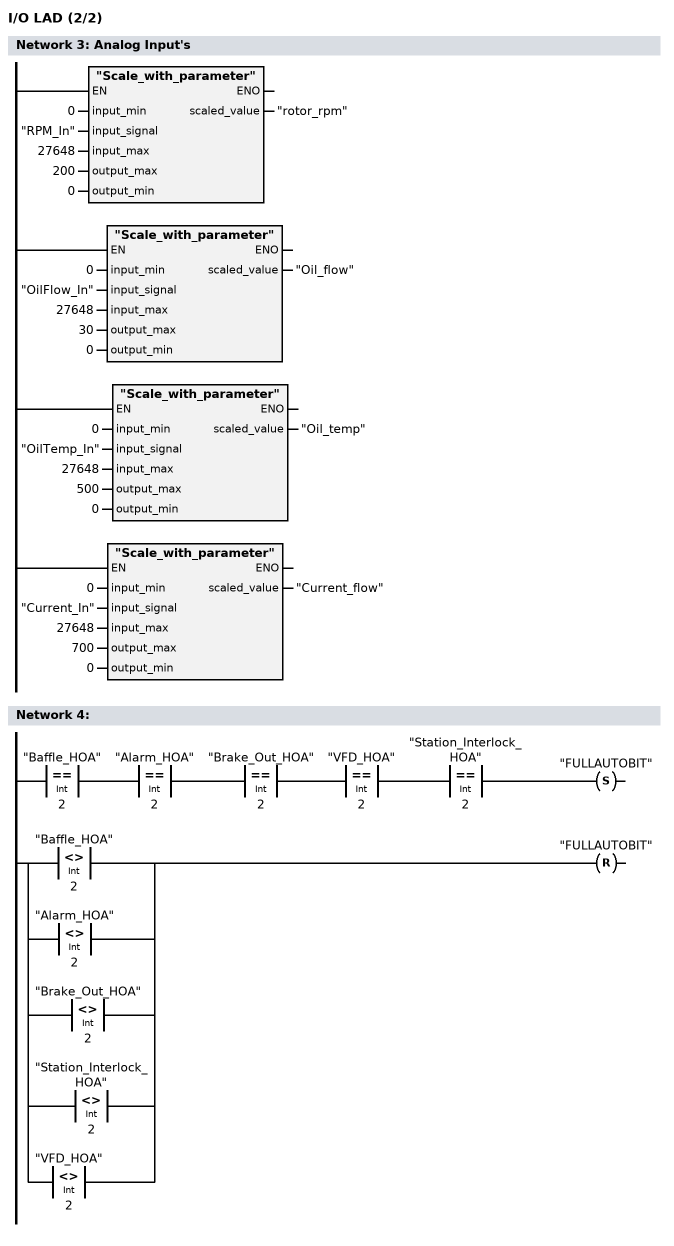
   RUNG wire#powerrail
      "Scale_with_parameter"(input_min := 0, input_signal := "RPM_In", input_max := 27648, output_max := 200, output_min := 0, scaled_value => "rotor_rpm")
   END_RUNG
   RUNG wire#powerrail
      "Scale_with_parameter"(input_min := 0, input_signal := "OilFlow_In", input_max := 27648, output_max := 30, output_min := 0, scaled_value => "Oil_flow")
   END_RUNG
   RUNG wire#powerrail
      "Scale_with_parameter"(input_min := 0, input_signal := "OilTemp_In", input_max := 27648, output_max := 500, output_min := 0, scaled_value => "Oil_temp")
   END_RUNG
   RUNG wire#powerrail
      "Scale_with_parameter"(input_min := 0, input_signal := "Current_In", input_max := 27648, output_max := 700, output_min := 0, scaled_value => "Current_flow")
   END_RUNG
   // the same network as SCL:
   "Scale_with_parameter"(input_min := 0,
                          input_signal := "RPM_In",
                          input_max := 27648,
                          output_max := 200,
                          output_min := 0,
                          scaled_value => "rotor_rpm");
   "Scale_with_parameter"(input_min := 0,
                          input_signal := "OilFlow_In",
                          input_max := 27648,
                          output_max := 30,
                          output_min := 0,
                          scaled_value => "Oil_flow");
   "Scale_with_parameter"(input_min := 0,
                          input_signal := "OilTemp_In",
                          input_max := 27648,
                          output_max := 500,
                          output_min := 0,
                          scaled_value => "Oil_temp");
   "Scale_with_parameter"(input_min := 0,
                          input_signal := "Current_In",
                          input_max := 27648,
                          output_max := 700,
                          output_min := 0,
                          scaled_value => "Current_flow");
END_REGION

REGION Network 4
   RUNG wire#powerrail
      { S7_Templates := "SrcType := Int" } EQ_Contact(in1 := "Baffle_HOA", in2 := 2)
      { S7_Templates := "SrcType := Int" } EQ_Contact(in1 := "Alarm_HOA", in2 := 2)
      { S7_Templates := "SrcType := Int" } EQ_Contact(in1 := "Brake_Out_HOA", in2 := 2)
      { S7_Templates := "SrcType := Int" } EQ_Contact(in1 := "VFD_HOA", in2 := 2)
      { S7_Templates := "SrcType := Int" } EQ_Contact(in1 := "Station_Interlock_HOA", in2 := 2)
      S_Coil( "FULLAUTOBIT" )
   END_RUNG
   RUNG wire#powerrail
      { S7_Templates := "SrcType := Int" } NE_Contact(in1 := "Baffle_HOA", in2 := 2)
      wire#w1
      R_Coil( "FULLAUTOBIT" )
   END_RUNG
   RUNG wire#powerrail
      { S7_Templates := "SrcType := Int" } NE_Contact(in1 := "Alarm_HOA", in2 := 2)
   END_RUNG wire#w1
   RUNG wire#powerrail
      { S7_Templates := "SrcType := Int" } NE_Contact(in1 := "Brake_Out_HOA", in2 := 2)
   END_RUNG wire#w1
   RUNG wire#powerrail
      { S7_Templates := "SrcType := Int" } NE_Contact(in1 := "Station_Interlock_HOA", in2 := 2)
   END_RUNG wire#w1
   RUNG wire#powerrail
      { S7_Templates := "SrcType := Int" } NE_Contact(in1 := "VFD_HOA", in2 := 2)
   END_RUNG wire#w1
   // the same network as SCL:
   IF ("Baffle_HOA" = 2) AND ("Alarm_HOA" = 2) AND ("Brake_Out_HOA" = 2) AND ("VFD_HOA" = 2) AND ("Station_Interlock_HOA" = 2) THEN
       "FULLAUTOBIT" := TRUE;
   END_IF;
   IF ("Baffle_HOA" <> 2) OR ("Alarm_HOA" <> 2) OR ("Brake_Out_HOA" <> 2) OR ("Station_Interlock_HOA" <> 2) OR ("VFD_HOA" <> 2) THEN
       "FULLAUTOBIT" := FALSE;
   END_IF;
END_REGION
END_FUNCTION_BLOCK

FUNCTION_BLOCK "HOA_LAD"   // FB6, LAD
TITLE = Push Button for HOA (OFF, HAND, AUTO)
{ S7_Optimized_Access := 'TRUE' }
VERSION : 0.1
   VAR
      Os3 : Bool;
      Os2 : Bool;
      Os1 : Bool;
      Os4 : Bool;
      Os5 : Bool;
      Os6 : Bool;
      Os7 : Bool;
      Os8 : Bool;
      Os9 : Bool;
      Os10 : Bool;
      Os11 : Bool;
      Os12 : Bool;
   END_VAR
   VAR_TEMP   // added for the SCL form of the ladder/FBD networks
      _w1 : Bool;
      _w2 : Bool;
      _w3 : Bool;
   END_VAR
BEGIN

REGION Network 1
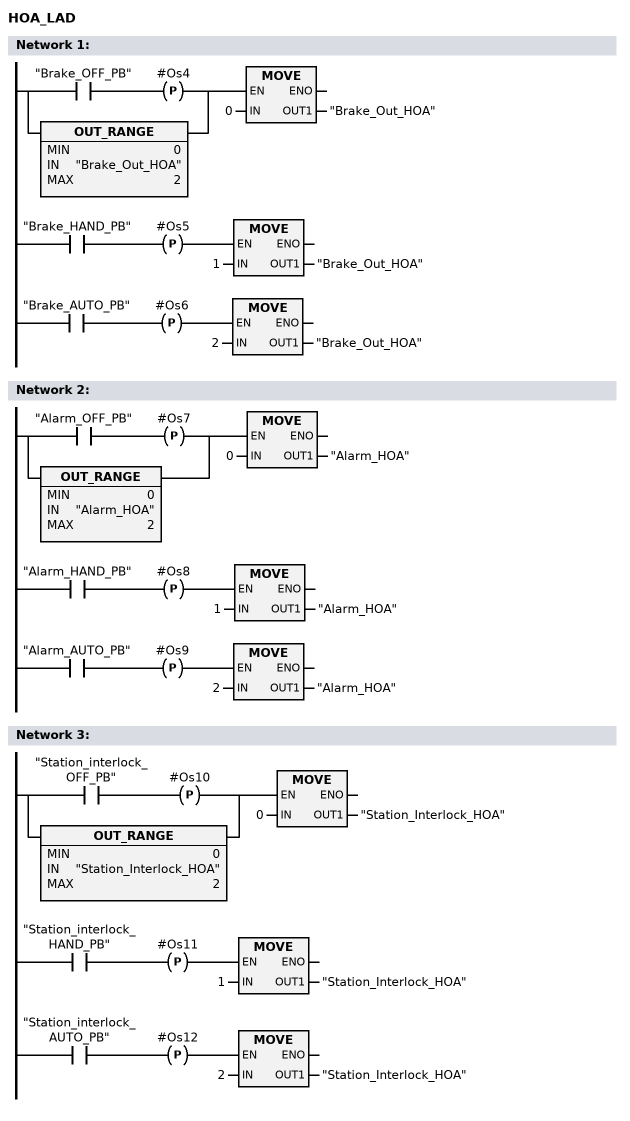
   #_w1 := "Brake_OFF_PB" AND NOT #Os4;   // rising edge
   #Os4 := "Brake_OFF_PB";
   IF #_w1 OR ("Brake_Out_HOA" < 0) OR ("Brake_Out_HOA" > 2) THEN "Brake_Out_HOA" := 0; END_IF;
   #_w2 := "Brake_HAND_PB" AND NOT #Os5;   // rising edge
   #Os5 := "Brake_HAND_PB";
   IF #_w2 THEN "Brake_Out_HOA" := 1; END_IF;
   #_w3 := "Brake_AUTO_PB" AND NOT #Os6;   // rising edge
   #Os6 := "Brake_AUTO_PB";
   IF #_w3 THEN "Brake_Out_HOA" := 2; END_IF;
END_REGION

REGION Network 2
   #_w1 := "Alarm_OFF_PB" AND NOT #Os7;   // rising edge
   #Os7 := "Alarm_OFF_PB";
   IF #_w1 OR ("Alarm_HOA" < 0) OR ("Alarm_HOA" > 2) THEN "Alarm_HOA" := 0; END_IF;
   #_w2 := "Alarm_HAND_PB" AND NOT #Os8;   // rising edge
   #Os8 := "Alarm_HAND_PB";
   IF #_w2 THEN "Alarm_HOA" := 1; END_IF;
   #_w3 := "Alarm_AUTO_PB" AND NOT #Os9;   // rising edge
   #Os9 := "Alarm_AUTO_PB";
   IF #_w3 THEN "Alarm_HOA" := 2; END_IF;
END_REGION

REGION Network 3
   #_w1 := "Station_interlock_OFF_PB" AND NOT #Os10;   // rising edge
   #Os10 := "Station_interlock_OFF_PB";
   IF #_w1 OR ("Station_Interlock_HOA" < 0) OR ("Station_Interlock_HOA" > 2) THEN
       "Station_Interlock_HOA" := 0;
   END_IF;
   #_w2 := "Station_interlock_HAND_PB" AND NOT #Os11;   // rising edge
   #Os11 := "Station_interlock_HAND_PB";
   IF #_w2 THEN "Station_Interlock_HOA" := 1; END_IF;
   #_w3 := "Station_interlock_AUTO_PB" AND NOT #Os12;   // rising edge
   #Os12 := "Station_interlock_AUTO_PB";
   IF #_w3 THEN "Station_Interlock_HOA" := 2; END_IF;
END_REGION
END_FUNCTION_BLOCK

FUNCTION_BLOCK "Alarm_LAD"   // FB10, LAD
{ S7_Optimized_Access := 'TRUE' }
VERSION : 0.1
   VAR
      OS1 : Bool;
      OS2 : Bool;
      OS3 : Bool;
      OS4 : Bool;
      OS5 : Bool;
      OS6 : Bool;
      OS7 : Bool;
      os8 : Bool;
   END_VAR
   VAR_TEMP
      tp1 : Int;
      OLFD : Time;
      OFL_AT : Bool;
      tp2 : Int;
      OCD : Time;
      OC_AT : Bool;
      tp3 : Int;
      HOT : Time;
      HOT_AT : Bool;
      tp4 : Int;
      ROS : Time;
      ROS_AT : Bool;
      tp5 : Int;
      OHF : Time;
      OHF_AT : Bool;
      tp6 : Int;
      BF : Time;
      BF_AT : Bool;
      ES_AT : Bool;
      AlarmTrigger : Bool;
   END_VAR
   VAR_TEMP   // added for the SCL form of the ladder/FBD networks
      _w1 : Bool;
      _w2 : Bool;
   END_VAR
BEGIN

REGION Network 1: Alarm for OIL LOW FLOW
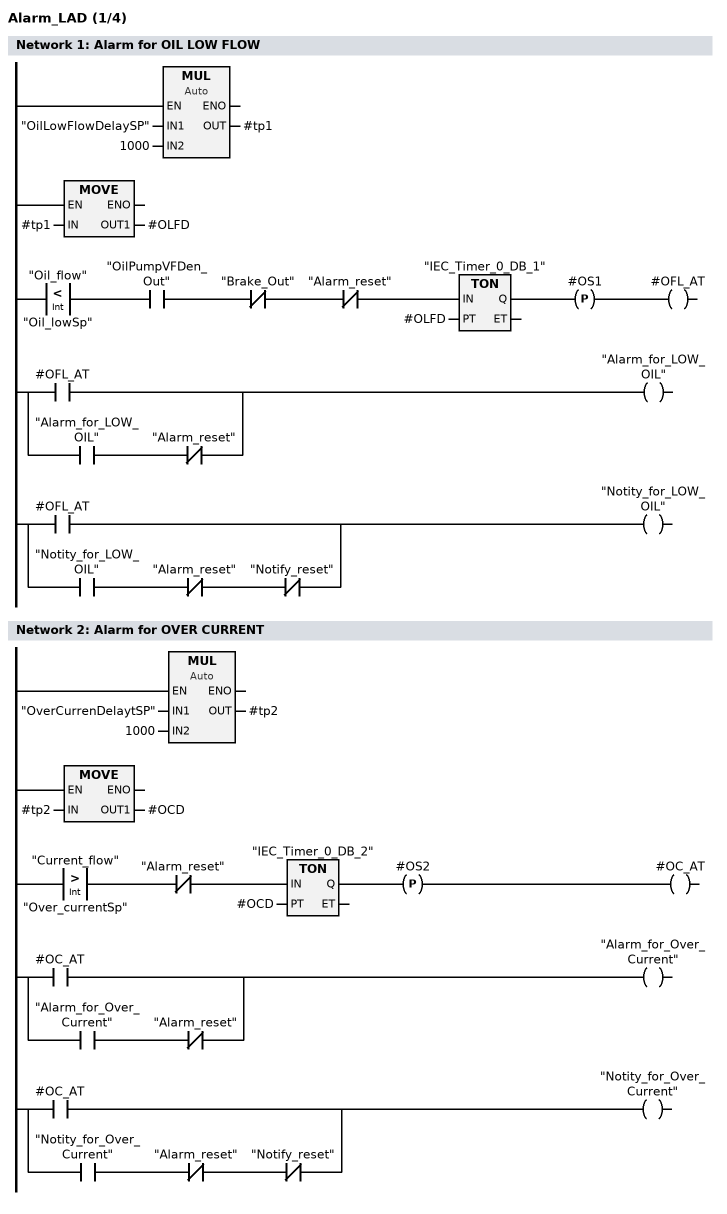
   #tp1 := "OilLowFlowDelaySP" * 1000;
   #OLFD := #tp1;
   "IEC_Timer_0_DB_1".TON(IN := ("Oil_flow" < "Oil_lowSp") AND "OilPumpVFDen_Out" AND NOT "Brake_Out" AND NOT "Alarm_reset",
                          PT := #OLFD);
   #_w1 := "IEC_Timer_0_DB_1".Q AND NOT #OS1;   // rising edge
   #OS1 := "IEC_Timer_0_DB_1".Q;
   #OFL_AT := #_w1;
   "Alarm_for_LOW_OIL" := #OFL_AT OR ("Alarm_for_LOW_OIL" AND NOT "Alarm_reset");
   "Notity_for_LOW_OIL" := #OFL_AT OR ("Notity_for_LOW_OIL" AND NOT "Alarm_reset" AND NOT "Notify_reset");
END_REGION

REGION Network 2: Alarm for OVER CURRENT
   #tp2 := "OverCurrenDelaytSP" * 1000;
   #OCD := #tp2;
   "IEC_Timer_0_DB_2".TON(IN := ("Current_flow" > "Over_currentSp") AND NOT "Alarm_reset", PT := #OCD);
   #_w1 := "IEC_Timer_0_DB_2".Q AND NOT #OS2;   // rising edge
   #OS2 := "IEC_Timer_0_DB_2".Q;
   #OC_AT := #_w1;
   "Alarm_for_Over_Current" := #OC_AT OR ("Alarm_for_Over_Current" AND NOT "Alarm_reset");
   "Notity_for_Over_Current" := #OC_AT OR ("Notity_for_Over_Current" AND NOT "Alarm_reset" AND NOT "Notify_reset");
END_REGION

REGION Network 3: Alarm for High Oil Temp
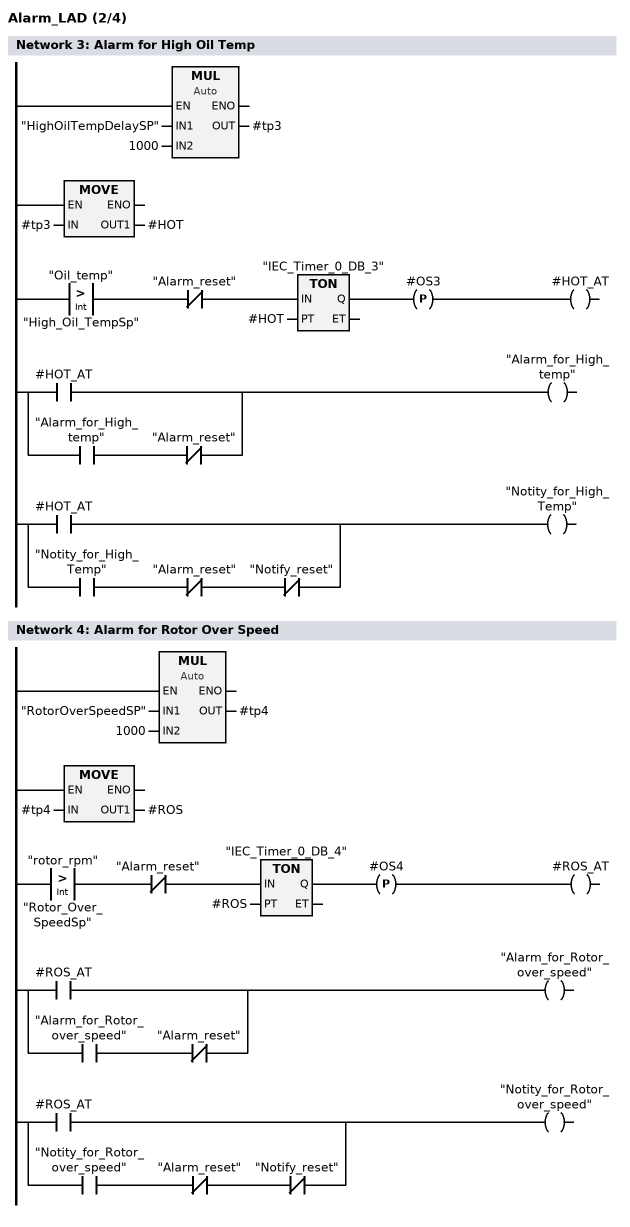
   #tp3 := "HighOilTempDelaySP" * 1000;
   #HOT := #tp3;
   "IEC_Timer_0_DB_3".TON(IN := ("Oil_temp" > "High_Oil_TempSp") AND NOT "Alarm_reset", PT := #HOT);
   #_w1 := "IEC_Timer_0_DB_3".Q AND NOT #OS3;   // rising edge
   #OS3 := "IEC_Timer_0_DB_3".Q;
   #HOT_AT := #_w1;
   "Alarm_for_High_temp" := #HOT_AT OR ("Alarm_for_High_temp" AND NOT "Alarm_reset");
   "Notity_for_High_Temp" := #HOT_AT OR ("Notity_for_High_Temp" AND NOT "Alarm_reset" AND NOT "Notify_reset");
END_REGION

REGION Network 4: Alarm for Rotor Over Speed
   #tp4 := "RotorOverSpeedSP" * 1000;
   #ROS := #tp4;
   "IEC_Timer_0_DB_4".TON(IN := ("rotor_rpm" > "Rotor_Over_SpeedSp") AND NOT "Alarm_reset", PT := #ROS);
   #_w1 := "IEC_Timer_0_DB_4".Q AND NOT #OS4;   // rising edge
   #OS4 := "IEC_Timer_0_DB_4".Q;
   #ROS_AT := #_w1;
   "Alarm_for_Rotor_over_speed" := #ROS_AT OR ("Alarm_for_Rotor_over_speed" AND NOT "Alarm_reset");
   "Notity_for_Rotor_over_speed" := #ROS_AT OR ("Notity_for_Rotor_over_speed" AND NOT "Alarm_reset" AND NOT "Notify_reset");
END_REGION

REGION Network 5: Alarm for Oil High Flow
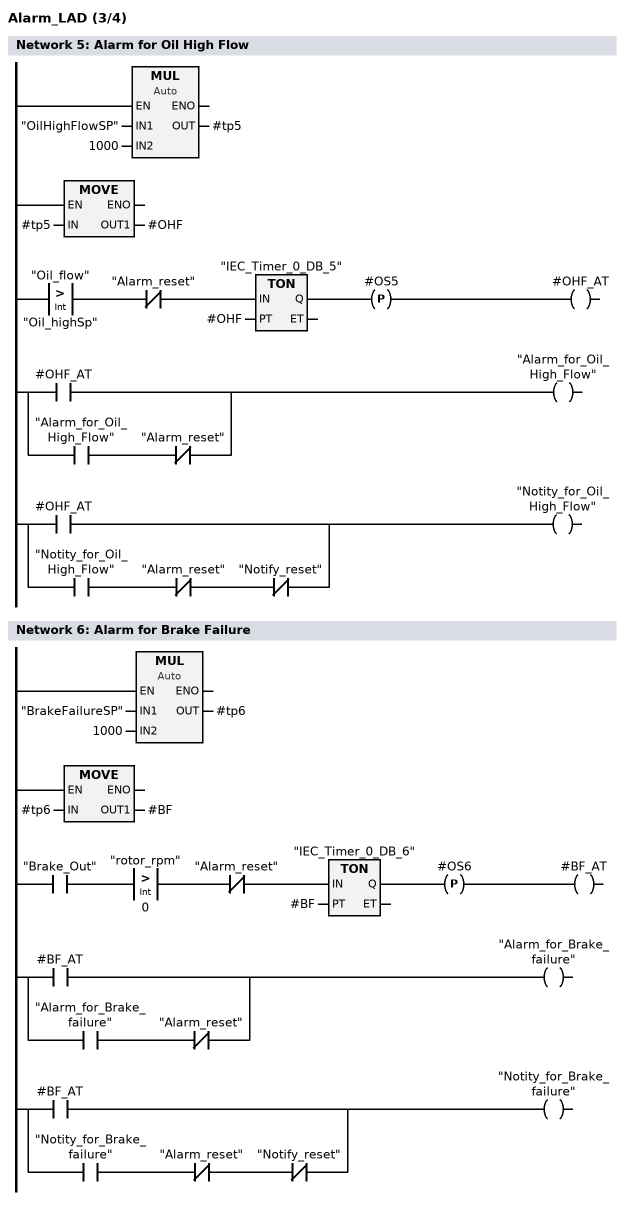
   #tp5 := "OilHighFlowSP" * 1000;
   #OHF := #tp5;
   "IEC_Timer_0_DB_5".TON(IN := ("Oil_flow" > "Oil_highSp") AND NOT "Alarm_reset", PT := #OHF);
   #_w1 := "IEC_Timer_0_DB_5".Q AND NOT #OS5;   // rising edge
   #OS5 := "IEC_Timer_0_DB_5".Q;
   #OHF_AT := #_w1;
   "Alarm_for_Oil_High_Flow" := #OHF_AT OR ("Alarm_for_Oil_High_Flow" AND NOT "Alarm_reset");
   "Notity_for_Oil_High_Flow" := #OHF_AT OR ("Notity_for_Oil_High_Flow" AND NOT "Alarm_reset" AND NOT "Notify_reset");
END_REGION

REGION Network 6: Alarm for Brake Failure
   #tp6 := "BrakeFailureSP" * 1000;
   #BF := #tp6;
   "IEC_Timer_0_DB_6".TON(IN := "Brake_Out" AND ("rotor_rpm" > 0) AND NOT "Alarm_reset", PT := #BF);
   #_w1 := "IEC_Timer_0_DB_6".Q AND NOT #OS6;   // rising edge
   #OS6 := "IEC_Timer_0_DB_6".Q;
   #BF_AT := #_w1;
   "Alarm_for_Brake_failure" := #BF_AT OR ("Alarm_for_Brake_failure" AND NOT "Alarm_reset");
   "Notity_for_Brake_failure" := #BF_AT OR ("Notity_for_Brake_failure" AND NOT "Alarm_reset" AND NOT "Notify_reset");
END_REGION

REGION Network 7: Alarm for E_STOP
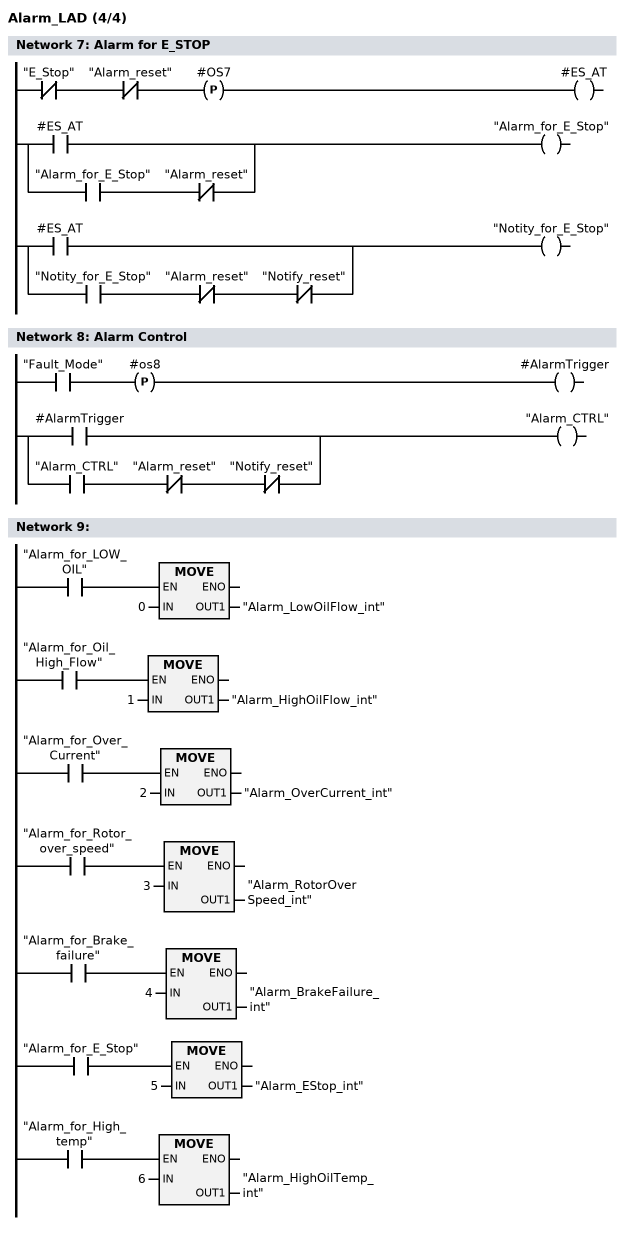
   RUNG wire#powerrail
      I_Contact( "E_Stop" )
      I_Contact( "Alarm_reset" )
      P_Trig( #OS7 )
      Coil( #ES_AT )
   END_RUNG
   RUNG wire#powerrail
      Contact( #ES_AT )
      wire#w1
      Coil( "Alarm_for_E_Stop" )
   END_RUNG
   RUNG wire#powerrail
      Contact( "Alarm_for_E_Stop" )
      I_Contact( "Alarm_reset" )
   END_RUNG wire#w1
   RUNG wire#powerrail
      Contact( #ES_AT )
      wire#w2
      Coil( "Notity_for_E_Stop" )
   END_RUNG
   RUNG wire#powerrail
      Contact( "Notity_for_E_Stop" )
      I_Contact( "Alarm_reset" )
      I_Contact( "Notify_reset" )
   END_RUNG wire#w2
   // the same network as SCL:
   #_w1 := NOT "E_Stop" AND NOT "Alarm_reset";
   #_w2 := #_w1 AND NOT #OS7;   // rising edge
   #OS7 := #_w1;
   #ES_AT := #_w2;
   "Alarm_for_E_Stop" := #ES_AT OR ("Alarm_for_E_Stop" AND NOT "Alarm_reset");
   "Notity_for_E_Stop" := #ES_AT OR ("Notity_for_E_Stop" AND NOT "Alarm_reset" AND NOT "Notify_reset");
END_REGION

REGION Network 8: Alarm Control
   RUNG wire#powerrail
      Contact( "Fault_Mode" )
      P_Trig( #os8 )
      Coil( #AlarmTrigger )
   END_RUNG
   RUNG wire#powerrail
      Contact( #AlarmTrigger )
      wire#w1
      Coil( "Alarm_CTRL" )
   END_RUNG
   RUNG wire#powerrail
      Contact( "Alarm_CTRL" )
      I_Contact( "Alarm_reset" )
      I_Contact( "Notify_reset" )
   END_RUNG wire#w1
   // the same network as SCL:
   #_w1 := "Fault_Mode" AND NOT #os8;   // rising edge
   #os8 := "Fault_Mode";
   #AlarmTrigger := #_w1;
   "Alarm_CTRL" := #AlarmTrigger OR ("Alarm_CTRL" AND NOT "Alarm_reset" AND NOT "Notify_reset");
END_REGION

REGION Network 9
   RUNG wire#powerrail
      Contact( "Alarm_for_LOW_OIL" )
      Move(in := 0, out1 => "Alarm_LowOilFlow_int")
   END_RUNG
   RUNG wire#powerrail
      Contact( "Alarm_for_Oil_High_Flow" )
      Move(in := 1, out1 => "Alarm_HighOilFlow_int")
   END_RUNG
   RUNG wire#powerrail
      Contact( "Alarm_for_Over_Current" )
      Move(in := 2, out1 => "Alarm_OverCurrent_int")
   END_RUNG
   RUNG wire#powerrail
      Contact( "Alarm_for_Rotor_over_speed" )
      Move(in := 3, out1 => "Alarm_RotorOverSpeed_int")
   END_RUNG
   RUNG wire#powerrail
      Contact( "Alarm_for_Brake_failure" )
      Move(in := 4, out1 => "Alarm_BrakeFailure_int")
   END_RUNG
   RUNG wire#powerrail
      Contact( "Alarm_for_E_Stop" )
      Move(in := 5, out1 => "Alarm_EStop_int")
   END_RUNG
   RUNG wire#powerrail
      Contact( "Alarm_for_High_temp" )
      Move(in := 6, out1 => "Alarm_HighOilTemp_int")
   END_RUNG
   // the same network as SCL:
   IF "Alarm_for_LOW_OIL" THEN "Alarm_LowOilFlow_int" := 0; END_IF;
   IF "Alarm_for_Oil_High_Flow" THEN "Alarm_HighOilFlow_int" := 1; END_IF;
   IF "Alarm_for_Over_Current" THEN "Alarm_OverCurrent_int" := 2; END_IF;
   IF "Alarm_for_Rotor_over_speed" THEN "Alarm_RotorOverSpeed_int" := 3; END_IF;
   IF "Alarm_for_Brake_failure" THEN "Alarm_BrakeFailure_int" := 4; END_IF;
   IF "Alarm_for_E_Stop" THEN "Alarm_EStop_int" := 5; END_IF;
   IF "Alarm_for_High_temp" THEN "Alarm_HighOilTemp_int" := 6; END_IF;
END_REGION
END_FUNCTION_BLOCK

FUNCTION_BLOCK "Modes_LAD"   // FB14, LAD
{ S7_Optimized_Access := 'TRUE' }
VERSION : 0.1
   VAR
      os1 : Bool;
      os2 : Bool;
      os3 : Bool;
      os4 : Bool;
      os5 : Bool;
   END_VAR
   VAR_TEMP
      tv1 : Int;
      ti1 : Time;
      tv3 : Int;
      tv2 : Int;
      tv4 : Int;
      ti2 : Time;
      tv5 : Int;
      ti3 : Time;
   END_VAR
   VAR_TEMP   // added for the SCL form of the ladder/FBD networks
      _w1 : Bool;
      _w2 : Bool;
      _w3 : Bool;
   END_VAR
BEGIN

REGION Network 1: WarmUp_Mode
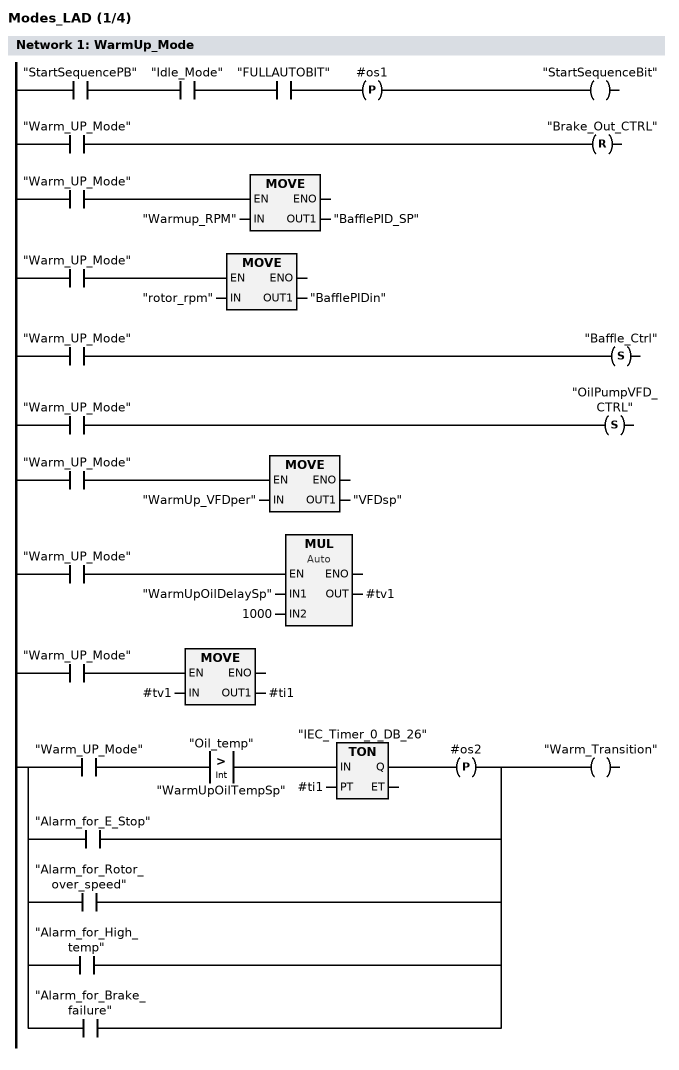
   #_w1 := "StartSequencePB" AND "Idle_Mode" AND "FULLAUTOBIT";
   #_w2 := #_w1 AND NOT #os1;   // rising edge
   #os1 := #_w1;
   "StartSequenceBit" := #_w2;
   IF "Warm_UP_Mode" THEN
       "Brake_Out_CTRL" := FALSE;
       "BafflePID_SP" := "Warmup_RPM";
       "BafflePIDin" := "rotor_rpm";
       "Baffle_Ctrl" := TRUE;
       "OilPumpVFD_CTRL" := TRUE;
       "VFDsp" := "WarmUp_VFDper";
       #tv1 := "WarmUpOilDelaySp" * 1000;
       #ti1 := #tv1;
   END_IF;
   "IEC_Timer_0_DB_26".TON(IN := "Warm_UP_Mode" AND ("Oil_temp" > "WarmUpOilTempSp"), PT := #ti1);
   #_w3 := "IEC_Timer_0_DB_26".Q AND NOT #os2;   // rising edge
   #os2 := "IEC_Timer_0_DB_26".Q;
   "Warm_Transition" := #_w3 OR "Alarm_for_E_Stop" OR "Alarm_for_Rotor_over_speed" OR "Alarm_for_High_temp" OR "Alarm_for_Brake_failure";
END_REGION

REGION Network 2: Stabilize Mode
   // Generator should speed up until desired kW output is attained. Once we’re stable within 
   // 5kW (+/-) of the setpoint for at least 10 seconds, we should transition into the next mode.
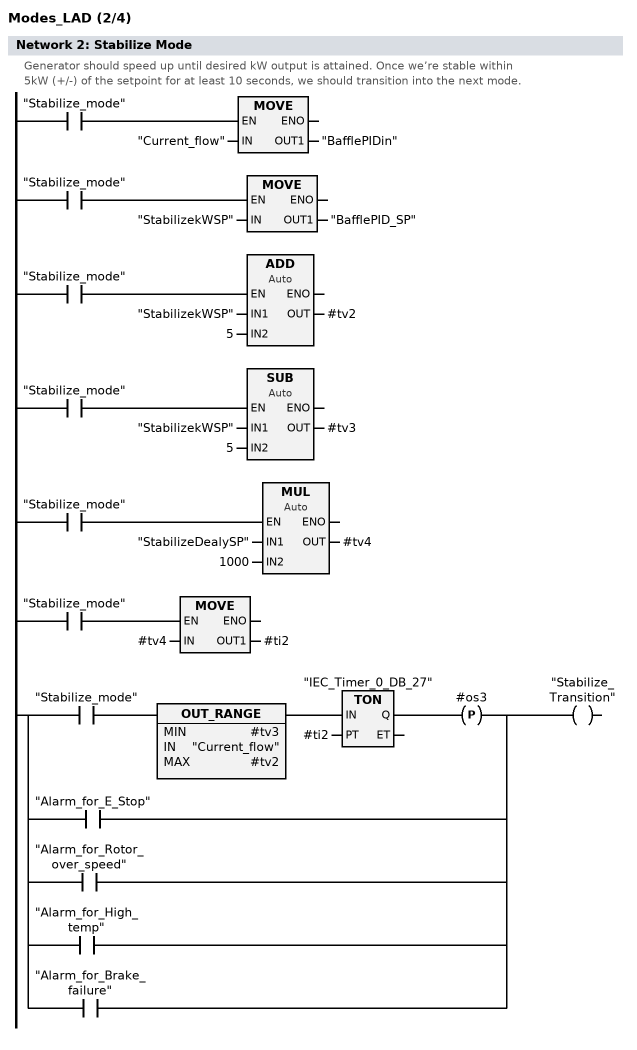
   IF "Stabilize_mode" THEN
       "BafflePIDin" := "Current_flow";
       "BafflePID_SP" := "StabilizekWSP";
       #tv2 := "StabilizekWSP" + 5;
       #tv3 := "StabilizekWSP" - 5;
       #tv4 := "StabilizeDealySP" * 1000;
       #ti2 := #tv4;
   END_IF;
   "IEC_Timer_0_DB_27".TON(IN := "Stabilize_mode" AND (("Current_flow" < #tv3) OR ("Current_flow" > #tv2)),
                           PT := #ti2);
   #_w1 := "IEC_Timer_0_DB_27".Q AND NOT #os3;   // rising edge
   #os3 := "IEC_Timer_0_DB_27".Q;
   "Stabilize_Transition" := #_w1 OR "Alarm_for_E_Stop" OR "Alarm_for_Rotor_over_speed" OR "Alarm_for_High_temp" OR "Alarm_for_Brake_failure";
END_REGION

REGION Network 3: Generation_Mode
   // Keep everything running and close the interlock.
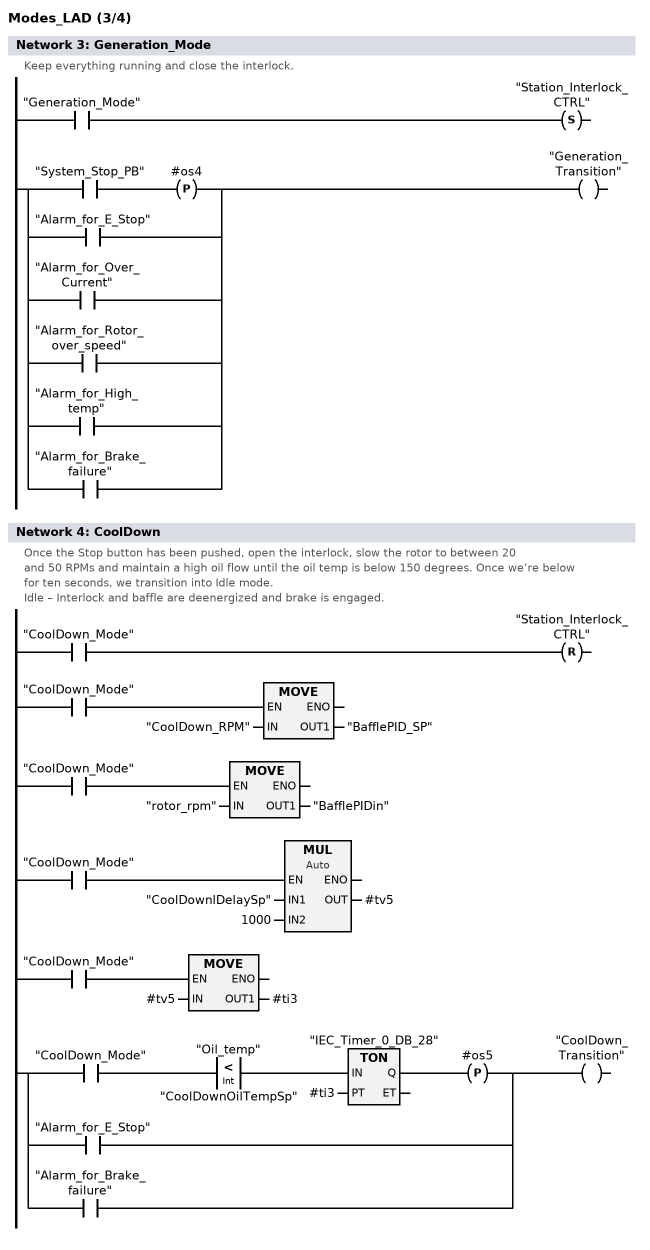
   RUNG wire#powerrail
      Contact( "Generation_Mode" )
      S_Coil( "Station_Interlock_CTRL" )
   END_RUNG
   RUNG wire#powerrail
      Contact( "System_Stop_PB" )
      P_Trig( #os4 )
      wire#w1
      Coil( "Generation_Transition" )
   END_RUNG
   RUNG wire#powerrail
      Contact( "Alarm_for_E_Stop" )
   END_RUNG wire#w1
   RUNG wire#powerrail
      Contact( "Alarm_for_Over_Current" )
   END_RUNG wire#w1
   RUNG wire#powerrail
      Contact( "Alarm_for_Rotor_over_speed" )
   END_RUNG wire#w1
   RUNG wire#powerrail
      Contact( "Alarm_for_High_temp" )
   END_RUNG wire#w1
   RUNG wire#powerrail
      Contact( "Alarm_for_Brake_failure" )
   END_RUNG wire#w1
   // the same network as SCL:
   IF "Generation_Mode" THEN "Station_Interlock_CTRL" := TRUE; END_IF;
   #_w1 := "System_Stop_PB" AND NOT #os4;   // rising edge
   #os4 := "System_Stop_PB";
   "Generation_Transition" := #_w1 OR "Alarm_for_E_Stop" OR "Alarm_for_Over_Current" OR "Alarm_for_Rotor_over_speed" OR "Alarm_for_High_temp" OR "Alarm_for_Brake_failure";
END_REGION

REGION Network 4: CoolDown
   // Once the Stop button has been pushed, open the interlock, slow the rotor to between 20 
   // and 50 RPMs and maintain a high oil flow until the oil temp is below 150 degrees. Once we’re below 
   // for ten seconds, we transition into Idle mode.
   //  Idle – Interlock and baffle are deenergized and brake is engaged.
   IF "CoolDown_Mode" THEN
       "Station_Interlock_CTRL" := FALSE;
       "BafflePID_SP" := "CoolDown_RPM";
       "BafflePIDin" := "rotor_rpm";
       #tv5 := "CoolDownlDelaySp" * 1000;
       #ti3 := #tv5;
   END_IF;
   "IEC_Timer_0_DB_28".TON(IN := "CoolDown_Mode" AND ("Oil_temp" < "CoolDownOilTempSp"), PT := #ti3);
   #_w1 := "IEC_Timer_0_DB_28".Q AND NOT #os5;   // rising edge
   #os5 := "IEC_Timer_0_DB_28".Q;
   "CoolDown_Transition" := #_w1 OR "Alarm_for_E_Stop" OR "Alarm_for_Brake_failure";
END_REGION

REGION Network 5: Idle Mode
   // Idle – Interlock and baffle are deenergized and brake is engaged.
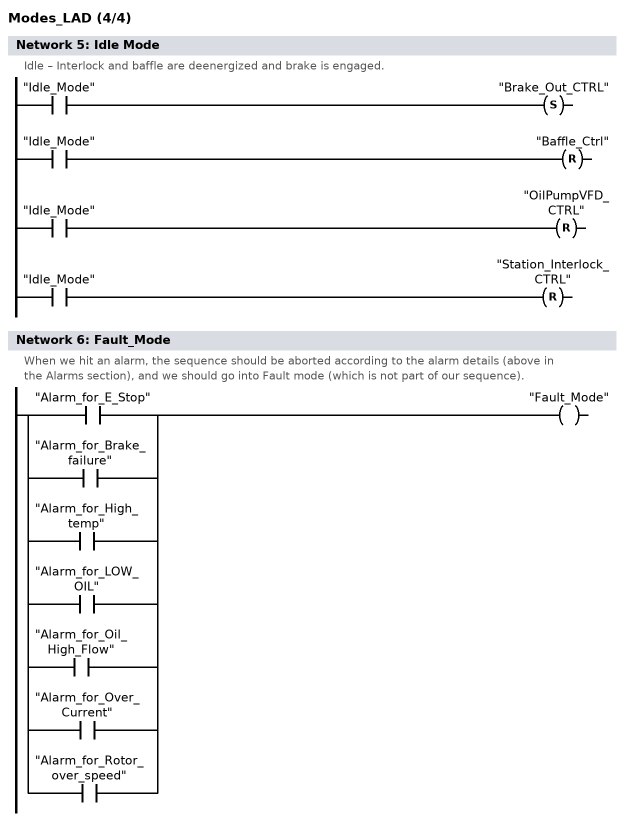
   RUNG wire#powerrail
      Contact( "Idle_Mode" )
      S_Coil( "Brake_Out_CTRL" )
   END_RUNG
   RUNG wire#powerrail
      Contact( "Idle_Mode" )
      R_Coil( "Baffle_Ctrl" )
   END_RUNG
   RUNG wire#powerrail
      Contact( "Idle_Mode" )
      R_Coil( "OilPumpVFD_CTRL" )
   END_RUNG
   RUNG wire#powerrail
      Contact( "Idle_Mode" )
      R_Coil( "Station_Interlock_CTRL" )
   END_RUNG
   // the same network as SCL:
   IF "Idle_Mode" THEN
       "Brake_Out_CTRL" := TRUE;
       "Baffle_Ctrl" := FALSE;
       "OilPumpVFD_CTRL" := FALSE;
       "Station_Interlock_CTRL" := FALSE;
   END_IF;
END_REGION
